(* Logix 5000 project; controller PLC_MCC1300_75F1 vendor 1 type 14 code 166 rev 32.11; software revision 32.04; part 48 of 83 *)
(* tags used below, declared in another part *)
   CONST_rgdDestMask : DINT[32];   // Destination Mask
   CONST_tPlant : UDT_PLANT_CONSTANTS;
   GP_TrackingSearchPlate : GP_TrackingSearchPlate;
   GP_TrackingValidateIndex : GP_TrackingValidateIndex;
   M30xTrimDeck_HMR : MAC_TrimmingDeck_HMR[5];
   M30xTrimWheel : MAC_TrimmingWheels[5];
   M30xTrimWheel_HMR : MAC_TrimmingWheels_HMR[5];
   M30xTrimWheel_HMW : MAC_TrimmingWheels_HMW[5];
   TMP_d : DINT;
   TMP_dHalfWidthDifference : DINT;
   TMP_dIndex : DINT;
   TMP_dMaskAllowed : DINT;
   TMP_xAllLiteToCullet : BOOL;
   TMP_xAtLeastOneForQuality : BOOL;
   TMP_xAtLeastOneForSideLeg : BOOL;
   TMP_xAtLeastOneOK : BOOL;
   xAlwaysOFF : BOOL;
   Z300_BufferPlate : UDT_LINE_BUFFER_PLATE;
   Z300_LineTracking : UDT_LINE_TRACKING;
(* MainProgram, continued *)

ROUTINE M30xTrimWheelBrManagement   (* ladder *)
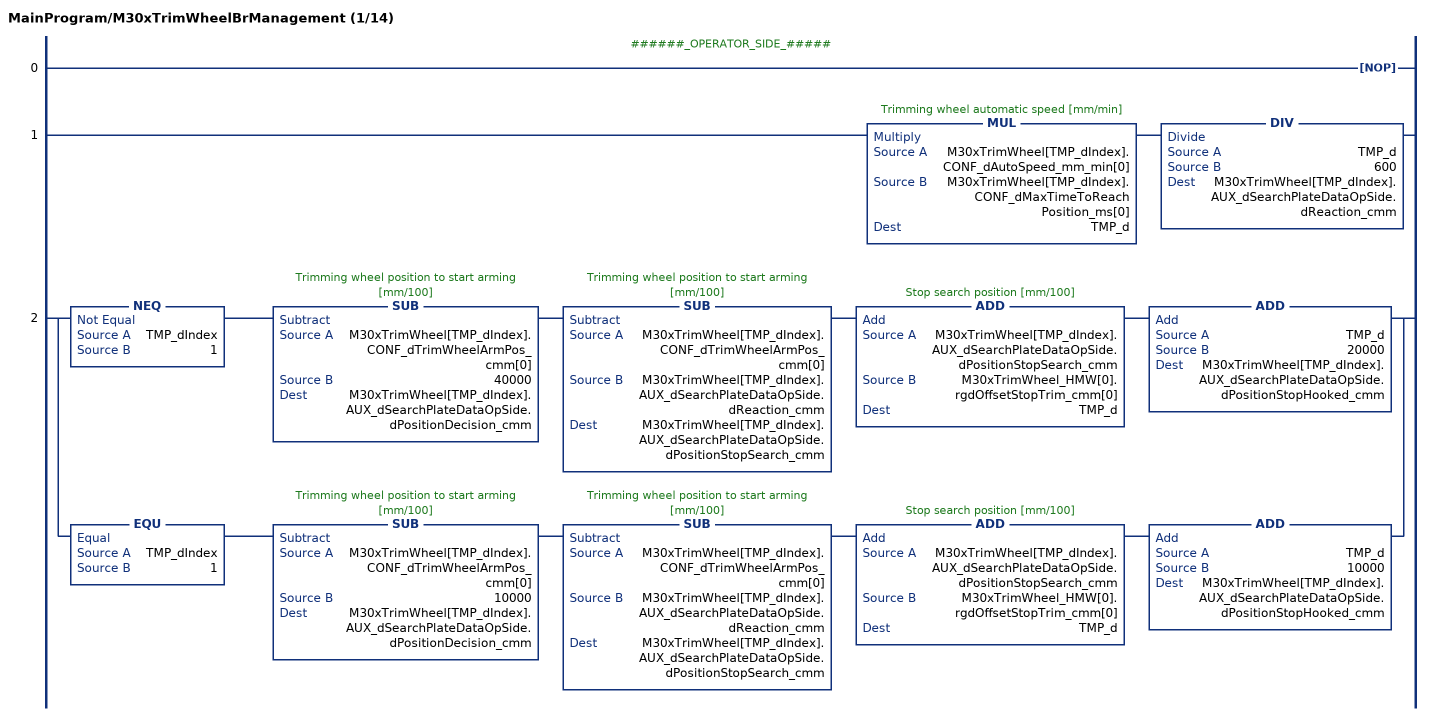
   // ######_OPERATOR_SIDE_#####
   0: NOP();
   1: MUL(M30xTrimWheel[TMP_dIndex].CONF_dAutoSpeed_mm_min[0],M30xTrimWheel[TMP_dIndex].CONF_dMaxTimeToReachPosition_ms[0],TMP_d)DIV(TMP_d,600,M30xTrimWheel[TMP_dIndex].AUX_dSearchPlateDataOpSide.dReaction_cmm);
   2: [NEQ(TMP_dIndex,1) SUB(M30xTrimWheel[TMP_dIndex].CONF_dTrimWheelArmPos_cmm[0],40000,M30xTrimWheel[TMP_dIndex].AUX_dSearchPlateDataOpSide.dPositionDecision_cmm) SUB(M30xTrimWheel[TMP_dIndex].CONF_dTrimWheelArmPos_cmm[0],M30xTrimWheel[TMP_dIndex].AUX_dSearchPlateDataOpSide.dReaction_cmm,M30xTrimWheel[TMP_dIndex].AUX_dSearchPlateDataOpSide.dPositionStopSearch_cmm) ADD(M30xTrimWheel[TMP_dIndex].AUX_dSearchPlateDataOpSide.dPositionStopSearch_cmm,M30xTrimWheel_HMW[0].rgdOffsetStopTrim_cmm[0],TMP_d) ADD(TMP_d,20000,M30xTrimWheel[TMP_dIndex].AUX_dSearchPlateDataOpSide.dPositionStopHooked_cmm) ,EQU(TMP_dIndex,1) SUB(M30xTrimWheel[TMP_dIndex].CONF_dTrimWheelArmPos_cmm[0],10000,M30xTrimWheel[TMP_dIndex].AUX_dSearchPlateDataOpSide.dPositionDecision_cmm) SUB(M30xTrimWheel[TMP_dIndex].CONF_dTrimWheelArmPos_cmm[0],M30xTrimWheel[TMP_dIndex].AUX_dSearchPlateDataOpSide.dReaction_cmm,M30xTrimWheel[TMP_dIndex].AUX_dSearchPlateDataOpSide.dPositionStopSearch_cmm) ADD(M30xTrimWheel[TMP_dIndex].AUX_dSearchPlateDataOpSide.dPositionStopSearch_cmm,M30xTrimWheel_HMW[0].rgdOffsetStopTrim_cmm[0],TMP_d) ADD(TMP_d,10000,M30xTrimWheel[TMP_dIndex].AUX_dSearchPlateDataOpSide.dPositionStopHooked_cmm) ];
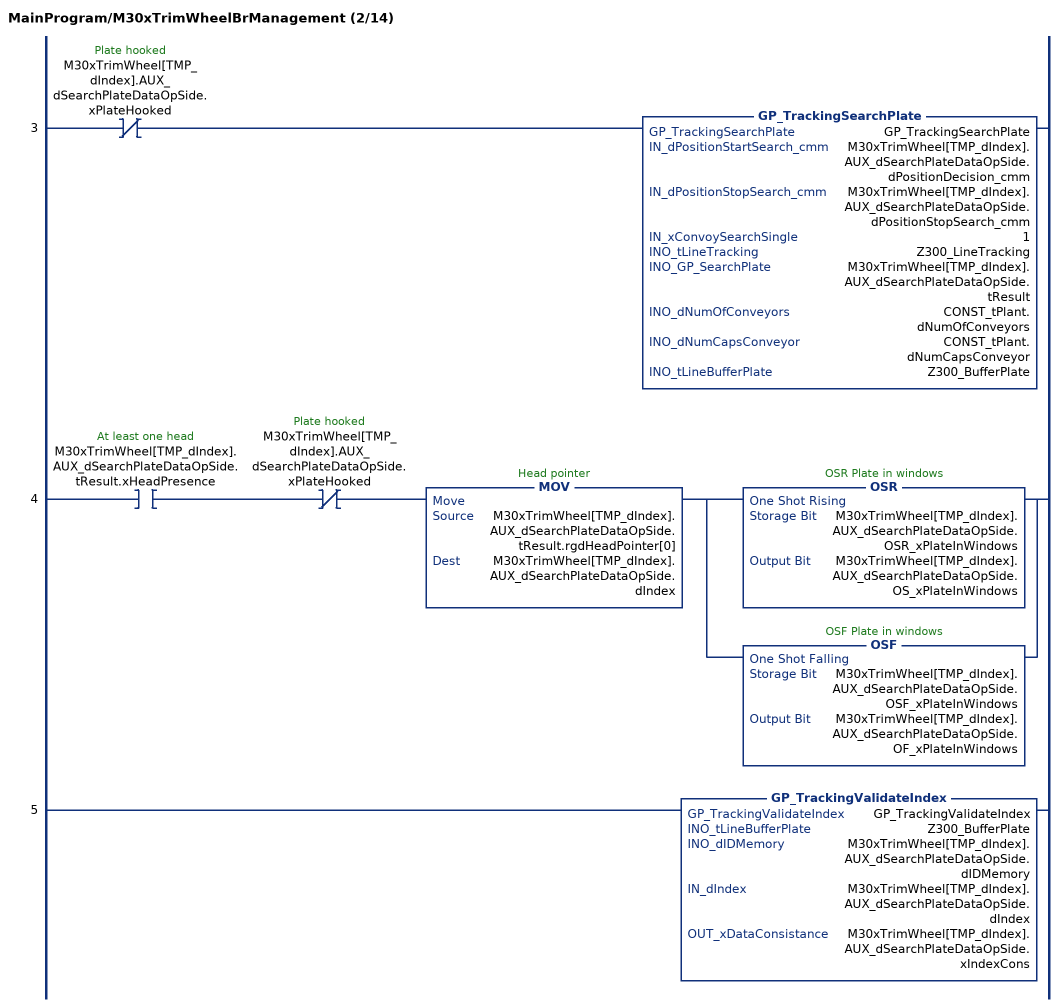
   3: XIO(M30xTrimWheel[TMP_dIndex].AUX_dSearchPlateDataOpSide.xPlateHooked)GP_TrackingSearchPlate(GP_TrackingSearchPlate,M30xTrimWheel[TMP_dIndex].AUX_dSearchPlateDataOpSide.dPositionDecision_cmm,M30xTrimWheel[TMP_dIndex].AUX_dSearchPlateDataOpSide.dPositionStopSearch_cmm,1,Z300_LineTracking,M30xTrimWheel[TMP_dIndex].AUX_dSearchPlateDataOpSide.tResult,CONST_tPlant.dNumOfConveyors,CONST_tPlant.dNumCapsConveyor,Z300_BufferPlate);
   4: XIC(M30xTrimWheel[TMP_dIndex].AUX_dSearchPlateDataOpSide.tResult.xHeadPresence)XIO(M30xTrimWheel[TMP_dIndex].AUX_dSearchPlateDataOpSide.xPlateHooked)MOV(M30xTrimWheel[TMP_dIndex].AUX_dSearchPlateDataOpSide.tResult.rgdHeadPointer[0],M30xTrimWheel[TMP_dIndex].AUX_dSearchPlateDataOpSide.dIndex)[OSR(M30xTrimWheel[TMP_dIndex].AUX_dSearchPlateDataOpSide.OSR_xPlateInWindows,M30xTrimWheel[TMP_dIndex].AUX_dSearchPlateDataOpSide.OS_xPlateInWindows) ,OSF(M30xTrimWheel[TMP_dIndex].AUX_dSearchPlateDataOpSide.OSF_xPlateInWindows,M30xTrimWheel[TMP_dIndex].AUX_dSearchPlateDataOpSide.OF_xPlateInWindows) ];
   5: GP_TrackingValidateIndex(GP_TrackingValidateIndex,Z300_BufferPlate,M30xTrimWheel[TMP_dIndex].AUX_dSearchPlateDataOpSide.dIDMemory,M30xTrimWheel[TMP_dIndex].AUX_dSearchPlateDataOpSide.dIndex,M30xTrimWheel[TMP_dIndex].AUX_dSearchPlateDataOpSide.xIndexCons);
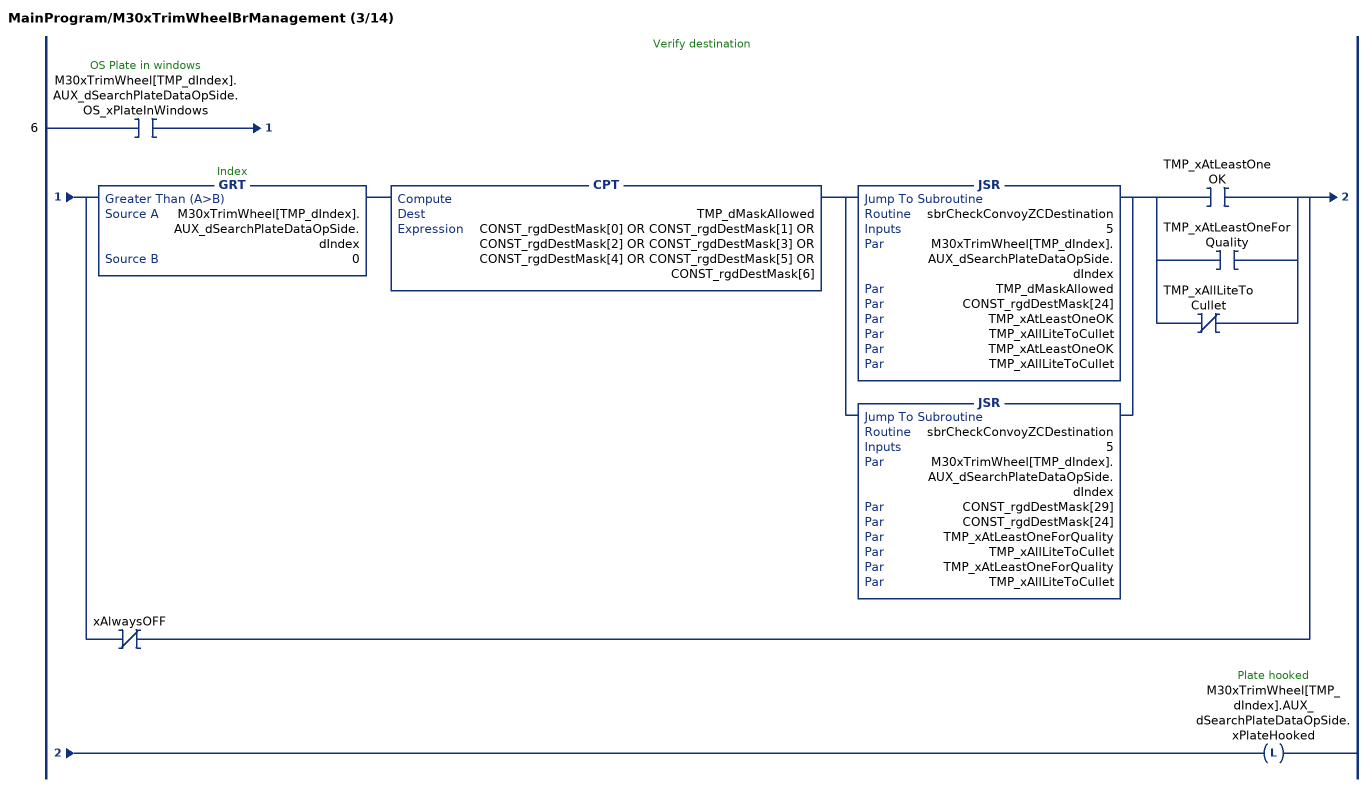
   // Verify destination
   6: XIC(M30xTrimWheel[TMP_dIndex].AUX_dSearchPlateDataOpSide.OS_xPlateInWindows)[GRT(M30xTrimWheel[TMP_dIndex].AUX_dSearchPlateDataOpSide.dIndex,0) CPT(TMP_dMaskAllowed,CONST_rgdDestMask[0] OR CONST_rgdDestMask[1] OR CONST_rgdDestMask[2] OR CONST_rgdDestMask[3] OR CONST_rgdDestMask[4] OR CONST_rgdDestMask[5] OR CONST_rgdDestMask[6]) [JSR(sbrCheckConvoyZCDestination,5,M30xTrimWheel[TMP_dIndex].AUX_dSearchPlateDataOpSide.dIndex,TMP_dMaskAllowed,CONST_rgdDestMask[24],TMP_xAtLeastOneOK,TMP_xAllLiteToCullet,TMP_xAtLeastOneOK,TMP_xAllLiteToCullet) ,JSR(sbrCheckConvoyZCDestination,5,M30xTrimWheel[TMP_dIndex].AUX_dSearchPlateDataOpSide.dIndex,CONST_rgdDestMask[29],CONST_rgdDestMask[24],TMP_xAtLeastOneForQuality,TMP_xAllLiteToCullet,TMP_xAtLeastOneForQuality,TMP_xAllLiteToCullet) ] [XIC(TMP_xAtLeastOneOK) ,XIC(TMP_xAtLeastOneForQuality) ,XIO(TMP_xAllLiteToCullet) ] ,XIO(xAlwaysOFF) ]OTL(M30xTrimWheel[TMP_dIndex].AUX_dSearchPlateDataOpSide.xPlateHooked);
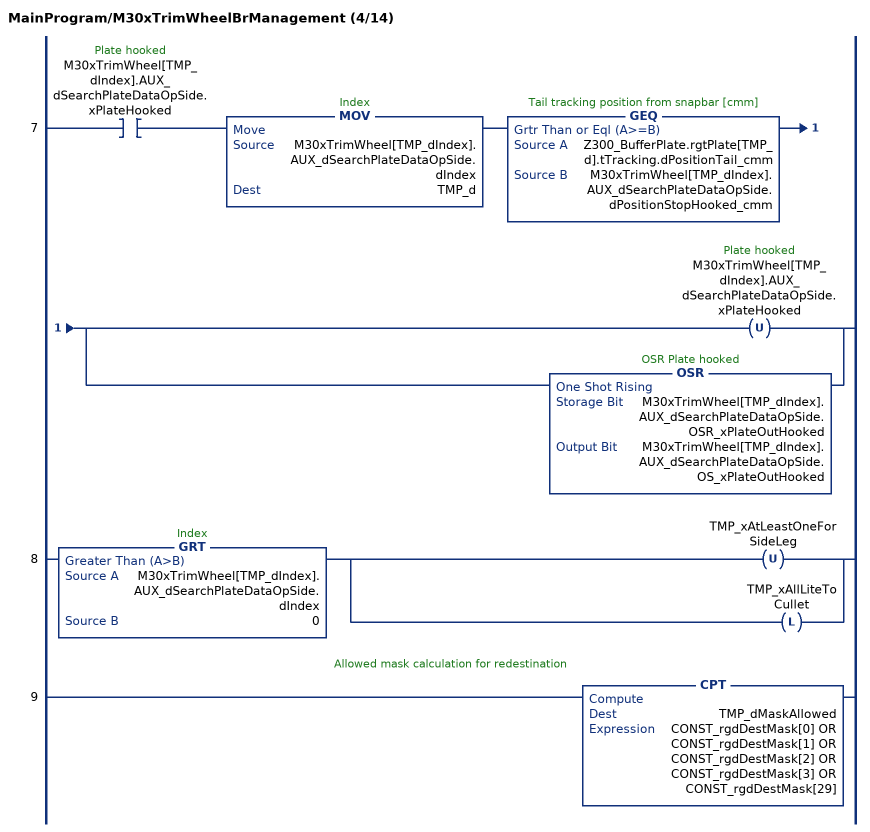
   7: XIC(M30xTrimWheel[TMP_dIndex].AUX_dSearchPlateDataOpSide.xPlateHooked)MOV(M30xTrimWheel[TMP_dIndex].AUX_dSearchPlateDataOpSide.dIndex,TMP_d)GEQ(Z300_BufferPlate.rgtPlate[TMP_d].tTracking.dPositionTail_cmm,M30xTrimWheel[TMP_dIndex].AUX_dSearchPlateDataOpSide.dPositionStopHooked_cmm)[OTU(M30xTrimWheel[TMP_dIndex].AUX_dSearchPlateDataOpSide.xPlateHooked) ,OSR(M30xTrimWheel[TMP_dIndex].AUX_dSearchPlateDataOpSide.OSR_xPlateOutHooked,M30xTrimWheel[TMP_dIndex].AUX_dSearchPlateDataOpSide.OS_xPlateOutHooked) ];
   8: GRT(M30xTrimWheel[TMP_dIndex].AUX_dSearchPlateDataOpSide.dIndex,0)[OTU(TMP_xAtLeastOneForSideLeg) ,OTL(TMP_xAllLiteToCullet) ];
   // Allowed mask calculation for redestination
   9: CPT(TMP_dMaskAllowed,CONST_rgdDestMask[0] OR CONST_rgdDestMask[1] OR CONST_rgdDestMask[2] OR CONST_rgdDestMask[3] OR CONST_rgdDestMask[29]);
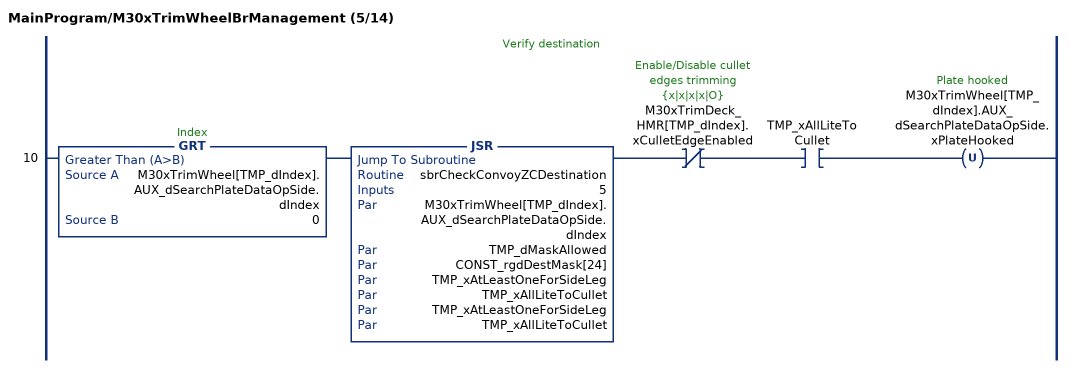
   // Verify destination
   10: GRT(M30xTrimWheel[TMP_dIndex].AUX_dSearchPlateDataOpSide.dIndex,0)JSR(sbrCheckConvoyZCDestination,5,M30xTrimWheel[TMP_dIndex].AUX_dSearchPlateDataOpSide.dIndex,TMP_dMaskAllowed,CONST_rgdDestMask[24],TMP_xAtLeastOneForSideLeg,TMP_xAllLiteToCullet,TMP_xAtLeastOneForSideLeg,TMP_xAllLiteToCullet)XIO(M30xTrimDeck_HMR[TMP_dIndex].xCulletEdgeEnabled)XIC(TMP_xAllLiteToCullet)OTU(M30xTrimWheel[TMP_dIndex].AUX_dSearchPlateDataOpSide.xPlateHooked);
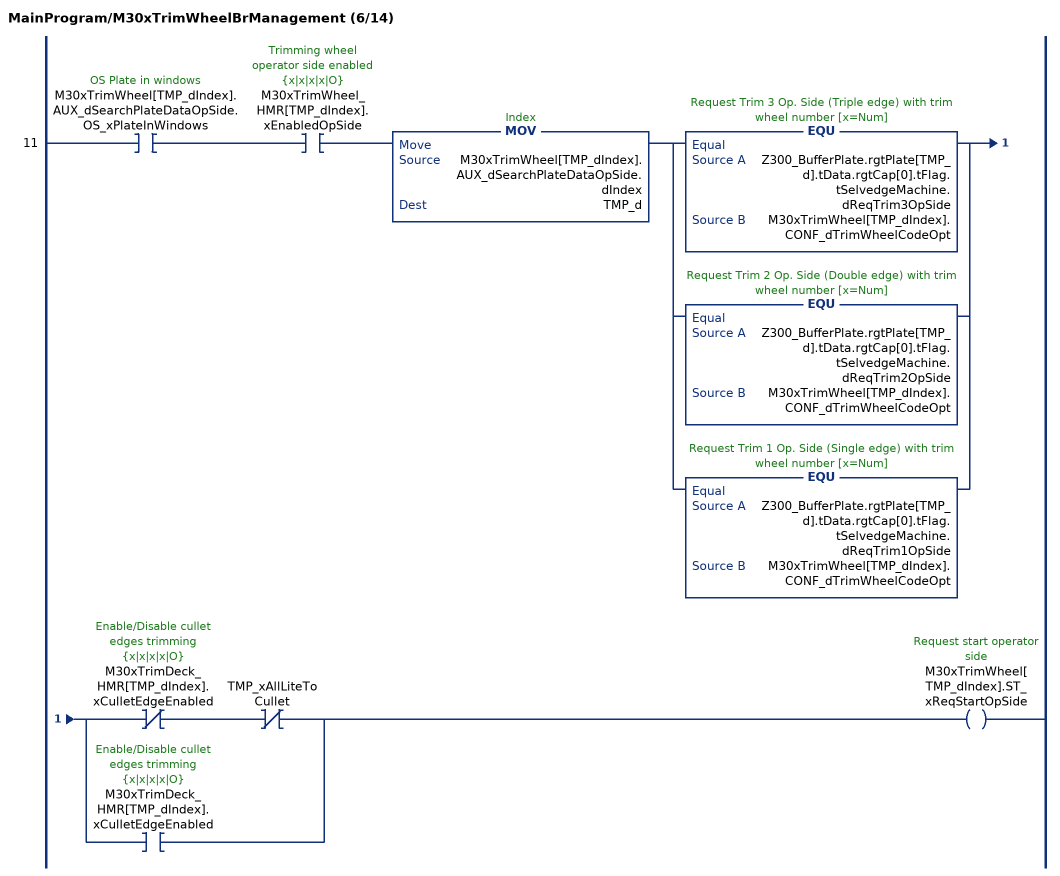
   11: XIC(M30xTrimWheel[TMP_dIndex].AUX_dSearchPlateDataOpSide.OS_xPlateInWindows)XIC(M30xTrimWheel_HMR[TMP_dIndex].xEnabledOpSide)MOV(M30xTrimWheel[TMP_dIndex].AUX_dSearchPlateDataOpSide.dIndex,TMP_d)[EQU(Z300_BufferPlate.rgtPlate[TMP_d].tData.rgtCap[0].tFlag.tSelvedgeMachine.dReqTrim3OpSide,M30xTrimWheel[TMP_dIndex].CONF_dTrimWheelCodeOpt) ,EQU(Z300_BufferPlate.rgtPlate[TMP_d].tData.rgtCap[0].tFlag.tSelvedgeMachine.dReqTrim2OpSide,M30xTrimWheel[TMP_dIndex].CONF_dTrimWheelCodeOpt) ,EQU(Z300_BufferPlate.rgtPlate[TMP_d].tData.rgtCap[0].tFlag.tSelvedgeMachine.dReqTrim1OpSide,M30xTrimWheel[TMP_dIndex].CONF_dTrimWheelCodeOpt) ][XIO(M30xTrimDeck_HMR[TMP_dIndex].xCulletEdgeEnabled) XIO(TMP_xAllLiteToCullet) ,XIC(M30xTrimDeck_HMR[TMP_dIndex].xCulletEdgeEnabled) ]OTE(M30xTrimWheel[TMP_dIndex].ST_xReqStartOpSide);
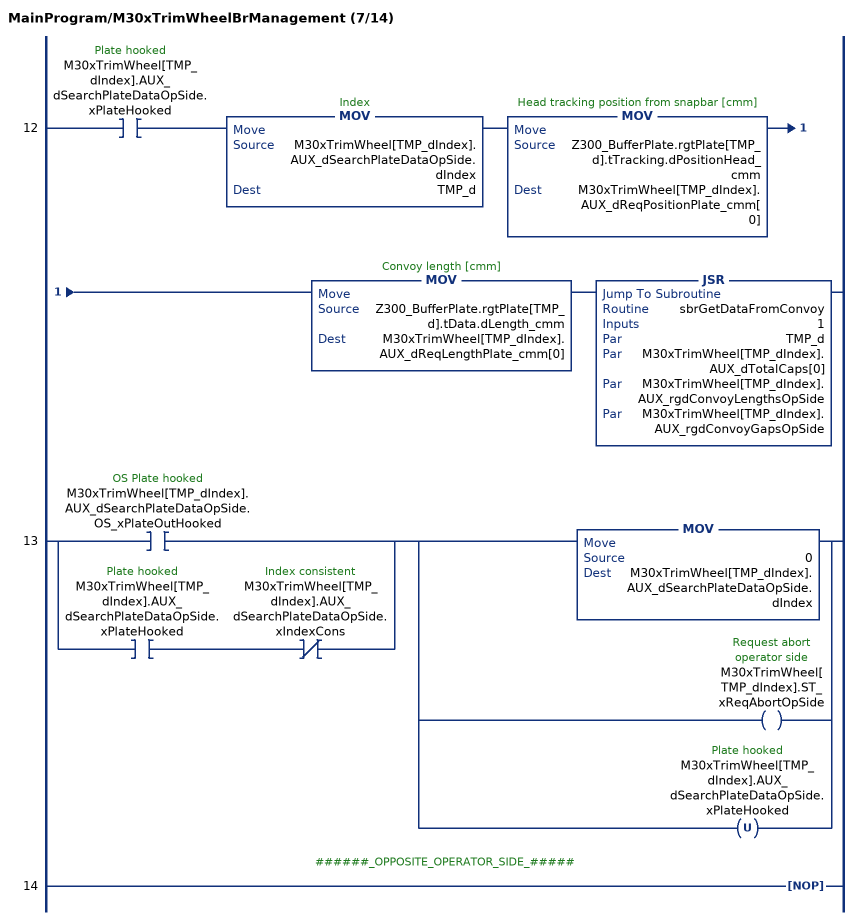
   12: XIC(M30xTrimWheel[TMP_dIndex].AUX_dSearchPlateDataOpSide.xPlateHooked)MOV(M30xTrimWheel[TMP_dIndex].AUX_dSearchPlateDataOpSide.dIndex,TMP_d)MOV(Z300_BufferPlate.rgtPlate[TMP_d].tTracking.dPositionHead_cmm,M30xTrimWheel[TMP_dIndex].AUX_dReqPositionPlate_cmm[0])MOV(Z300_BufferPlate.rgtPlate[TMP_d].tData.dLength_cmm,M30xTrimWheel[TMP_dIndex].AUX_dReqLengthPlate_cmm[0])JSR(sbrGetDataFromConvoy,1,TMP_d,M30xTrimWheel[TMP_dIndex].AUX_dTotalCaps[0],M30xTrimWheel[TMP_dIndex].AUX_rgdConvoyLengthsOpSide,M30xTrimWheel[TMP_dIndex].AUX_rgdConvoyGapsOpSide);
   13: [XIC(M30xTrimWheel[TMP_dIndex].AUX_dSearchPlateDataOpSide.OS_xPlateOutHooked) ,XIC(M30xTrimWheel[TMP_dIndex].AUX_dSearchPlateDataOpSide.xPlateHooked) XIO(M30xTrimWheel[TMP_dIndex].AUX_dSearchPlateDataOpSide.xIndexCons) ][MOV(0,M30xTrimWheel[TMP_dIndex].AUX_dSearchPlateDataOpSide.dIndex) ,OTE(M30xTrimWheel[TMP_dIndex].ST_xReqAbortOpSide) ,OTU(M30xTrimWheel[TMP_dIndex].AUX_dSearchPlateDataOpSide.xPlateHooked) ];
   // ######_OPPOSITE_OPERATOR_SIDE_#####
   14: NOP();
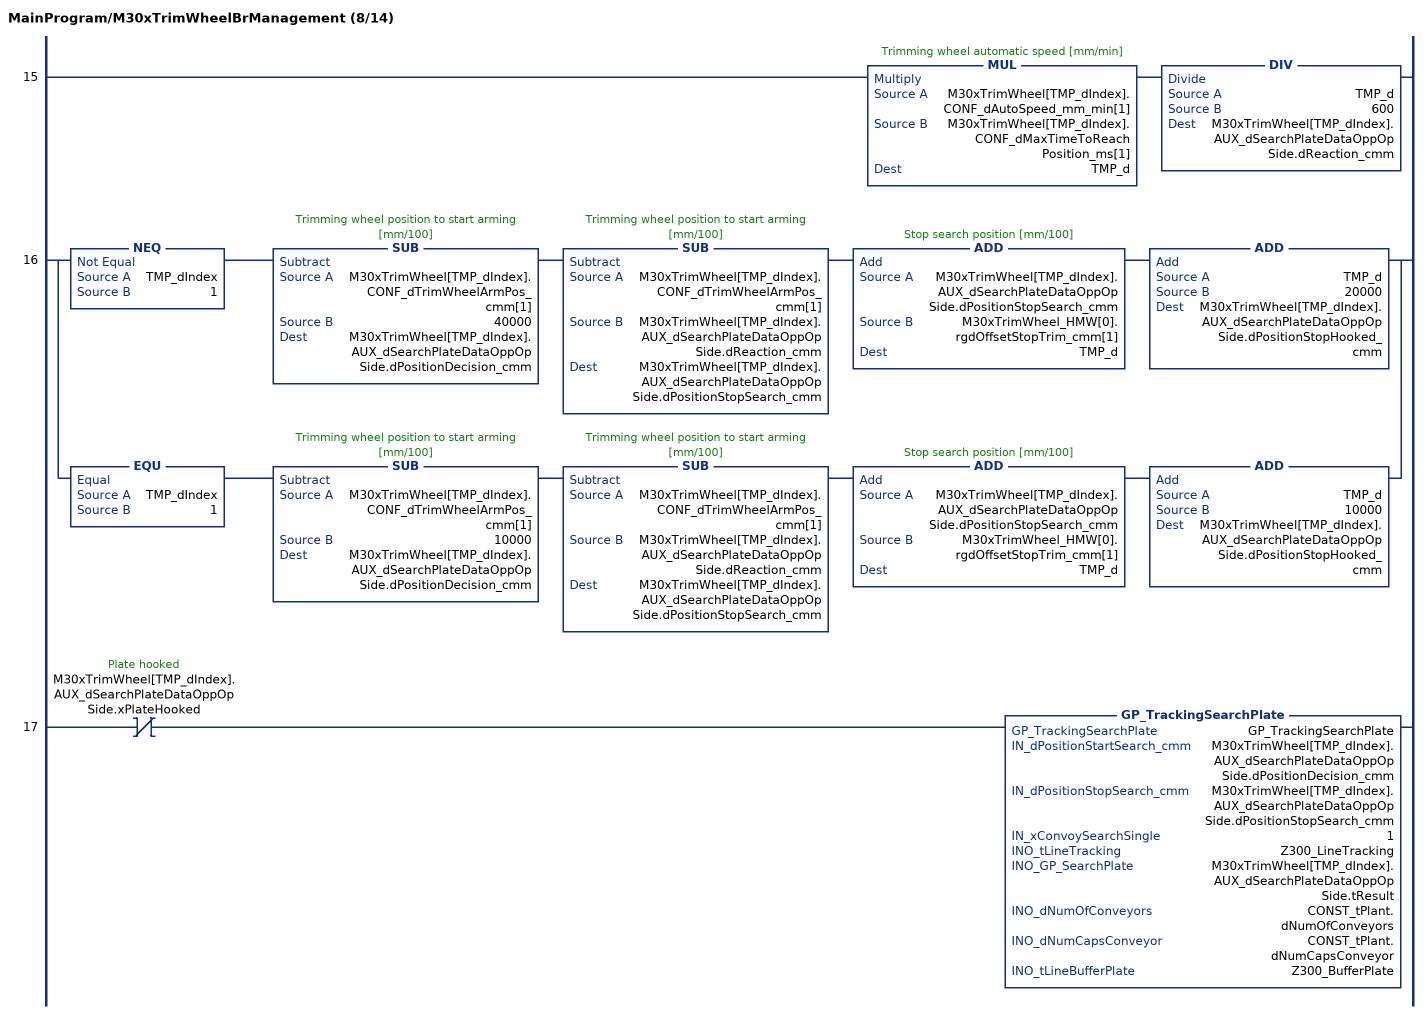
   15: MUL(M30xTrimWheel[TMP_dIndex].CONF_dAutoSpeed_mm_min[1],M30xTrimWheel[TMP_dIndex].CONF_dMaxTimeToReachPosition_ms[1],TMP_d)DIV(TMP_d,600,M30xTrimWheel[TMP_dIndex].AUX_dSearchPlateDataOppOpSide.dReaction_cmm);
   16: [NEQ(TMP_dIndex,1) SUB(M30xTrimWheel[TMP_dIndex].CONF_dTrimWheelArmPos_cmm[1],40000,M30xTrimWheel[TMP_dIndex].AUX_dSearchPlateDataOppOpSide.dPositionDecision_cmm) SUB(M30xTrimWheel[TMP_dIndex].CONF_dTrimWheelArmPos_cmm[1],M30xTrimWheel[TMP_dIndex].AUX_dSearchPlateDataOppOpSide.dReaction_cmm,M30xTrimWheel[TMP_dIndex].AUX_dSearchPlateDataOppOpSide.dPositionStopSearch_cmm) ADD(M30xTrimWheel[TMP_dIndex].AUX_dSearchPlateDataOppOpSide.dPositionStopSearch_cmm,M30xTrimWheel_HMW[0].rgdOffsetStopTrim_cmm[1],TMP_d) ADD(TMP_d,20000,M30xTrimWheel[TMP_dIndex].AUX_dSearchPlateDataOppOpSide.dPositionStopHooked_cmm) ,EQU(TMP_dIndex,1) SUB(M30xTrimWheel[TMP_dIndex].CONF_dTrimWheelArmPos_cmm[1],10000,M30xTrimWheel[TMP_dIndex].AUX_dSearchPlateDataOppOpSide.dPositionDecision_cmm) SUB(M30xTrimWheel[TMP_dIndex].CONF_dTrimWheelArmPos_cmm[1],M30xTrimWheel[TMP_dIndex].AUX_dSearchPlateDataOppOpSide.dReaction_cmm,M30xTrimWheel[TMP_dIndex].AUX_dSearchPlateDataOppOpSide.dPositionStopSearch_cmm) ADD(M30xTrimWheel[TMP_dIndex].AUX_dSearchPlateDataOppOpSide.dPositionStopSearch_cmm,M30xTrimWheel_HMW[0].rgdOffsetStopTrim_cmm[1],TMP_d) ADD(TMP_d,10000,M30xTrimWheel[TMP_dIndex].AUX_dSearchPlateDataOppOpSide.dPositionStopHooked_cmm) ];
   17: XIO(M30xTrimWheel[TMP_dIndex].AUX_dSearchPlateDataOppOpSide.xPlateHooked)GP_TrackingSearchPlate(GP_TrackingSearchPlate,M30xTrimWheel[TMP_dIndex].AUX_dSearchPlateDataOppOpSide.dPositionDecision_cmm,M30xTrimWheel[TMP_dIndex].AUX_dSearchPlateDataOppOpSide.dPositionStopSearch_cmm,1,Z300_LineTracking,M30xTrimWheel[TMP_dIndex].AUX_dSearchPlateDataOppOpSide.tResult,CONST_tPlant.dNumOfConveyors,CONST_tPlant.dNumCapsConveyor,Z300_BufferPlate);
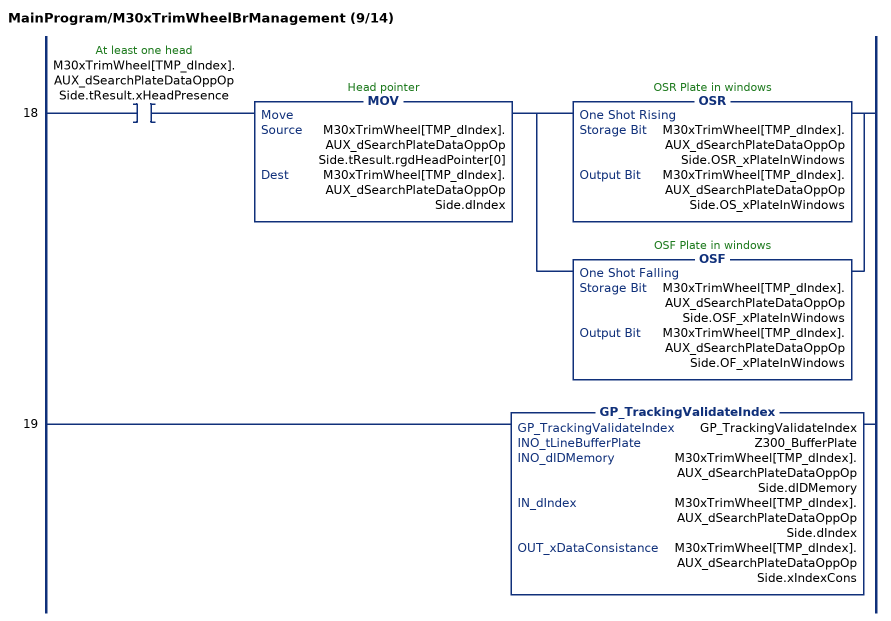
   18: XIC(M30xTrimWheel[TMP_dIndex].AUX_dSearchPlateDataOppOpSide.tResult.xHeadPresence)MOV(M30xTrimWheel[TMP_dIndex].AUX_dSearchPlateDataOppOpSide.tResult.rgdHeadPointer[0],M30xTrimWheel[TMP_dIndex].AUX_dSearchPlateDataOppOpSide.dIndex)[OSR(M30xTrimWheel[TMP_dIndex].AUX_dSearchPlateDataOppOpSide.OSR_xPlateInWindows,M30xTrimWheel[TMP_dIndex].AUX_dSearchPlateDataOppOpSide.OS_xPlateInWindows) ,OSF(M30xTrimWheel[TMP_dIndex].AUX_dSearchPlateDataOppOpSide.OSF_xPlateInWindows,M30xTrimWheel[TMP_dIndex].AUX_dSearchPlateDataOppOpSide.OF_xPlateInWindows) ];
   19: GP_TrackingValidateIndex(GP_TrackingValidateIndex,Z300_BufferPlate,M30xTrimWheel[TMP_dIndex].AUX_dSearchPlateDataOppOpSide.dIDMemory,M30xTrimWheel[TMP_dIndex].AUX_dSearchPlateDataOppOpSide.dIndex,M30xTrimWheel[TMP_dIndex].AUX_dSearchPlateDataOppOpSide.xIndexCons);
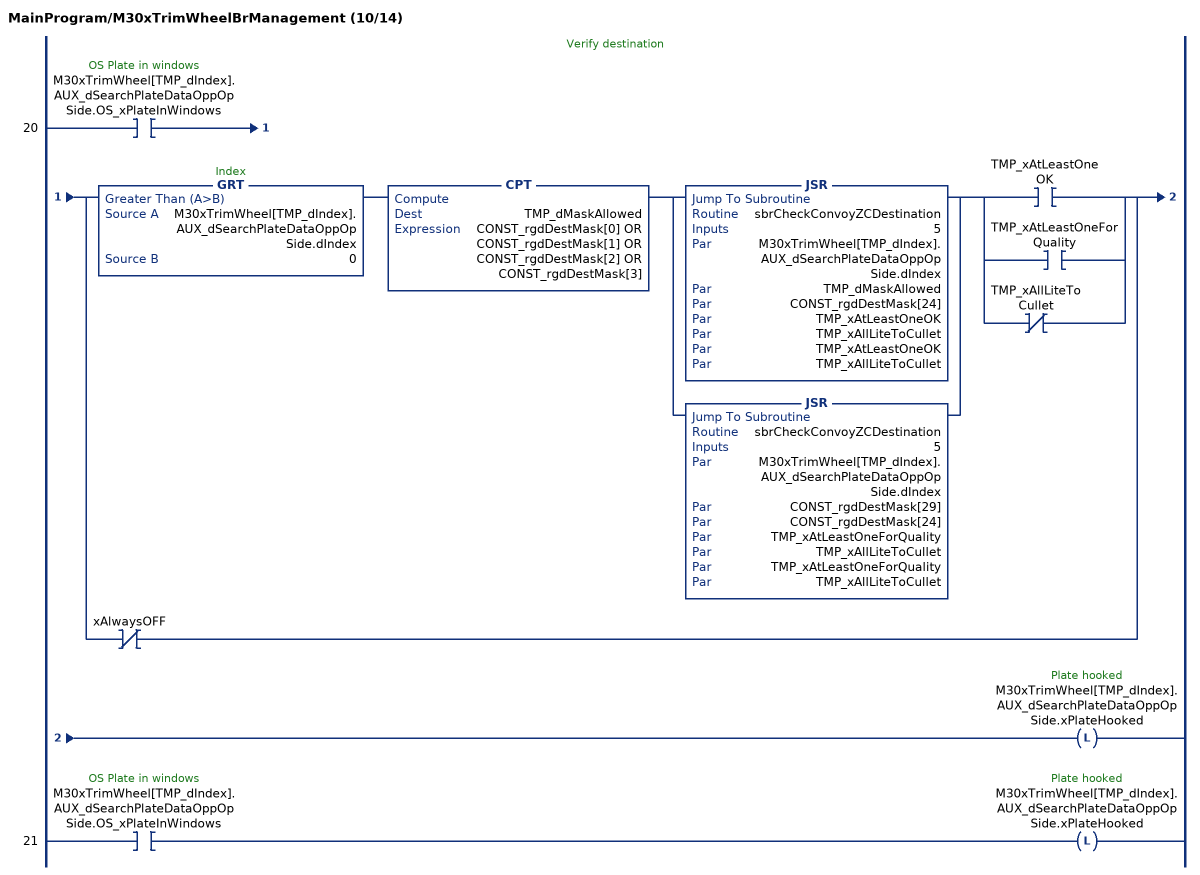
   // Verify destination
   20: XIC(M30xTrimWheel[TMP_dIndex].AUX_dSearchPlateDataOppOpSide.OS_xPlateInWindows)[GRT(M30xTrimWheel[TMP_dIndex].AUX_dSearchPlateDataOppOpSide.dIndex,0) CPT(TMP_dMaskAllowed,CONST_rgdDestMask[0] OR CONST_rgdDestMask[1] OR CONST_rgdDestMask[2] OR CONST_rgdDestMask[3]) [JSR(sbrCheckConvoyZCDestination,5,M30xTrimWheel[TMP_dIndex].AUX_dSearchPlateDataOppOpSide.dIndex,TMP_dMaskAllowed,CONST_rgdDestMask[24],TMP_xAtLeastOneOK,TMP_xAllLiteToCullet,TMP_xAtLeastOneOK,TMP_xAllLiteToCullet) ,JSR(sbrCheckConvoyZCDestination,5,M30xTrimWheel[TMP_dIndex].AUX_dSearchPlateDataOppOpSide.dIndex,CONST_rgdDestMask[29],CONST_rgdDestMask[24],TMP_xAtLeastOneForQuality,TMP_xAllLiteToCullet,TMP_xAtLeastOneForQuality,TMP_xAllLiteToCullet) ] [XIC(TMP_xAtLeastOneOK) ,XIC(TMP_xAtLeastOneForQuality) ,XIO(TMP_xAllLiteToCullet) ] ,XIO(xAlwaysOFF) ]OTL(M30xTrimWheel[TMP_dIndex].AUX_dSearchPlateDataOppOpSide.xPlateHooked);
   21: XIC(M30xTrimWheel[TMP_dIndex].AUX_dSearchPlateDataOppOpSide.OS_xPlateInWindows)OTL(M30xTrimWheel[TMP_dIndex].AUX_dSearchPlateDataOppOpSide.xPlateHooked);
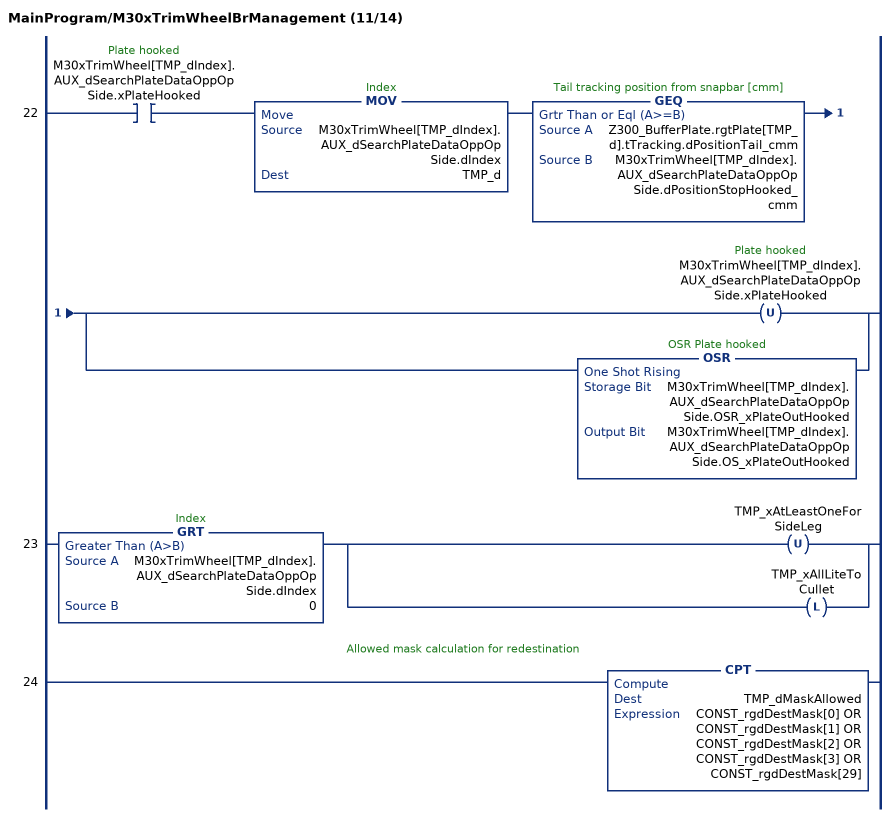
   22: XIC(M30xTrimWheel[TMP_dIndex].AUX_dSearchPlateDataOppOpSide.xPlateHooked)MOV(M30xTrimWheel[TMP_dIndex].AUX_dSearchPlateDataOppOpSide.dIndex,TMP_d)GEQ(Z300_BufferPlate.rgtPlate[TMP_d].tTracking.dPositionTail_cmm,M30xTrimWheel[TMP_dIndex].AUX_dSearchPlateDataOppOpSide.dPositionStopHooked_cmm)[OTU(M30xTrimWheel[TMP_dIndex].AUX_dSearchPlateDataOppOpSide.xPlateHooked) ,OSR(M30xTrimWheel[TMP_dIndex].AUX_dSearchPlateDataOppOpSide.OSR_xPlateOutHooked,M30xTrimWheel[TMP_dIndex].AUX_dSearchPlateDataOppOpSide.OS_xPlateOutHooked) ];
   23: GRT(M30xTrimWheel[TMP_dIndex].AUX_dSearchPlateDataOppOpSide.dIndex,0)[OTU(TMP_xAtLeastOneForSideLeg) ,OTL(TMP_xAllLiteToCullet) ];
   // Allowed mask calculation for redestination
   24: CPT(TMP_dMaskAllowed,CONST_rgdDestMask[0] OR CONST_rgdDestMask[1] OR CONST_rgdDestMask[2] OR CONST_rgdDestMask[3] OR CONST_rgdDestMask[29]);
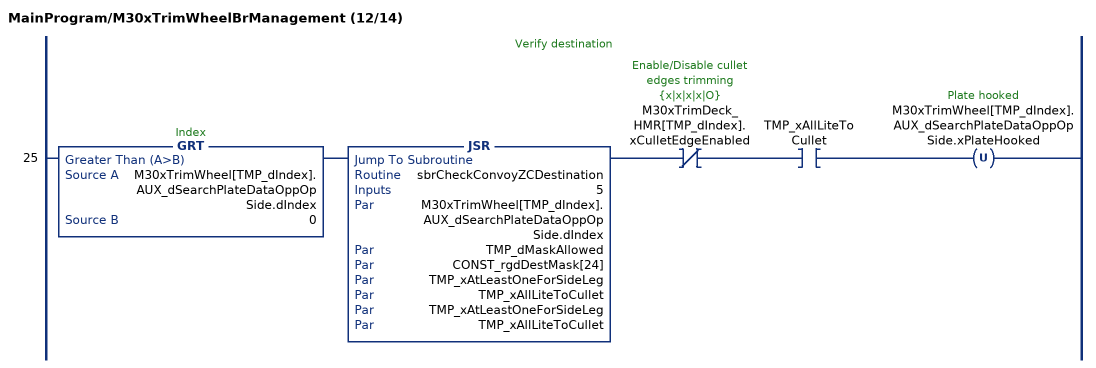
   // Verify destination
   25: GRT(M30xTrimWheel[TMP_dIndex].AUX_dSearchPlateDataOppOpSide.dIndex,0)JSR(sbrCheckConvoyZCDestination,5,M30xTrimWheel[TMP_dIndex].AUX_dSearchPlateDataOppOpSide.dIndex,TMP_dMaskAllowed,CONST_rgdDestMask[24],TMP_xAtLeastOneForSideLeg,TMP_xAllLiteToCullet,TMP_xAtLeastOneForSideLeg,TMP_xAllLiteToCullet)XIO(M30xTrimDeck_HMR[TMP_dIndex].xCulletEdgeEnabled)XIC(TMP_xAllLiteToCullet)OTU(M30xTrimWheel[TMP_dIndex].AUX_dSearchPlateDataOppOpSide.xPlateHooked);